
                       // FLAG information - store and evaluate
                       //------------------------------------------------------------------------------------------
                       // copy command setFlags for storing and usage in flag handling
                       // // setFlagsBuffer has twice the number of slots of PathDataPreBuffered to store flag information of past executed (already in MotionQueue) commands
                       #statFlagsBuffer.bufferElement[#statFlagsBuffer.writeBufferElement].pathDataName := #statPathDataPreBuffered.commands[#statPathDataPreBuffered.retrievePointer].pathDataName;
                       #statFlagsBuffer.bufferElement[#statFlagsBuffer.writeBufferElement].pathDataIdentifier := #statPathDataIdentifier;
                       #statFlagsBuffer.bufferElement[#statFlagsBuffer.writeBufferElement].cmdId := #statPathDataPreBuffered.commands[#statPathDataPreBuffered.retrievePointer].cmdID;
                       #statFlagsBuffer.bufferElement[#statFlagsBuffer.writeBufferElement].setFlags := #statPathDataPreBuffered.commands[#statPathDataPreBuffered.retrievePointer].setFlags;
                       #statFlagsBuffer.bufferElement[#statFlagsBuffer.writeBufferElement].valueFlags := #statPathDataPreBuffered.commands[#statPathDataPreBuffered.retrievePointer].valueFlags;
                       #statFlagsBuffer.bufferElement[#statFlagsBuffer.writeBufferElement].isIntermediateCmd := #statPathDataPreBuffered.commands[#statPathDataPreBuffered.retrievePointer].isIntermediateCmd;

                       // go to execution if cmd was copied
                       #statStateExecution := #EX_TRIGGERING_CMD;


                       IF #statPathDataPreBuffered.retrievePointer < "LKINCTRL_NO_OF_PATHDATA_PREBUFFER_ELEMENTS" THEN
                           #statPathDataPreBuffered.retrievePointer += 1;
                       ELSE
                           // restart PathDataPreBuf retrievePointer
                           #statPathDataPreBuffered.retrievePointer := 1;
                           // reset restart bit of pointer
                           #statPathDataPreBuffered.addPointerRestarted := FALSE;
                       END_IF;

                       #statSetFlagsBufferWriteBufferElement_old := #statFlagsBuffer.writeBufferElement;
                       // increase statSetFlagsBuffer write pointer and restart at overflow
                       IF #statFlagsBuffer.writeBufferElement < "LKINCTRL_NO_OF_SETFLAGS_BUFFER_ELEMENTS" THEN
                           #statFlagsBuffer.writeBufferElement := #statFlagsBuffer.writeBufferElement + 1;
                       ELSE
                           #statFlagsBuffer.writeBufferElement := 1;
                       END_IF;

                   ELSE
                       // set subfunction status according to PreBuffer status
                       IF (#statPathDataPreBuffered.retrievePointer = #statPathDataPreBuffered.addPointer
                           AND #statPathDataPreBuffered.addPointerRestarted = FALSE)
                       THEN
                           #statSubfunctionStatus := #STATUS_WAITING_FOR_PREBUFFERED_CMD;

                           // Check STOPRE signal from Parser/PreBuffer --> If true and executer is done then reset stopre to continue parsing
                           // PreBuffered commands are then executed and Parser and MovePath are in sync
                           IF #instLKinCtrl_MC_ExecuteKinMotionCmd.done AND #instLKinCtrl_PreBuffer.preprocessingStop THEN
                               #instLKinCtrl_PreBuffer.preprocessingStop := FALSE;
                           END_IF;


                       ELSIF (#statPathDataPreBuffered.addPointerRestarted = TRUE
                           AND (#statPathDataPreBuffered.retrievePointer - 1 = #statPathDataPreBuffered.addPointer))
                       THEN
                           #statSubfunctionStatus := #STATUS_PREBUFFERED_FULL;
                       END_IF;
                   END_IF;
                   // store old cmdID and PathDataName
                   #statPreBufferedCmdIdOld := #statPathDataElementPreBuffered.cmdID;
                   #statPreBufferedPathDataNameOld := #statPathDataElementPreBuffered.pathDataName;

                   // Check if interrupt was executed at start and if continue is needed
                   IF #statInterruptedAtStart THEN
                       IF #axesGroup.StatusMotionQueue.NumberOfCommands >= MIN(IN1:=#NO_OF_COMMANDS_PRELOADING, IN2:=#axesGroup.MotionQueue.MaxNumberOfCommands)
                           OR #statPathDataElementPreBuffered.cmdType = "LKINCTRL_CMD_WAIT_TIME" // Continue if waitTime shall be executed else we have deadlock
                           OR #statPathDataElementPreBuffered.cmdID = #statLastCmdIdPathdata // Continue if end of path was reached
                       THEN
                           #statStoreInterruptStateExecution := #statStateExecution;
                           #statStateExecution := #EX_CONTINUEING;
                           #statInterruptedAtStart := FALSE;
                       END_IF;
                   END_IF;

               END_IF;

           END_IF;
       END_REGION EX_GET_CMD


       // state reached when cmd should be triggered
       REGION EX_TRIGGERING_CMD
           IF #statStateExecution = #EX_TRIGGERING_CMD
               // AND #statDebugState = TRUE
               // wait condition bit (used for singleStep)
               AND #statExecutionWaitSingleStep = FALSE
               // wait condition bit (used for WAIT_TIME running)
               AND #statExecutionWaitTimerRunning = FALSE
               // wait condition bit (used for wait flags (acknowledge needed))
               AND #statWaitMain = FALSE
               // wait condition bit (used for wait value flags (acknowledge needed))
               AND #statWaitValueMain = FALSE
           THEN
               // reset  variable for single step debugging of states
               #statDebugState := FALSE;

               // call FB_ExecutePathMotion to execute cmd in same cycle
               #instLKinCtrl_MC_ExecuteKinMotionCmd(execute := TRUE,
                                                    interrupt := #interrupt,
                                                    stop := #stop,
                                                    pathDataElementPreBuf := #statPathDataElementPreBuffered,
                                                    conveyorConfiguration := #configuration.conveyorParameter,
                                                    to_Kinematics := #axesGroup);


               // check for cmd to be executed 
               IF #instLKinCtrl_MC_ExecuteKinMotionCmd.cmdExecuted THEN
                   // evaluate flag information for wait flags
                   // check for cmdId not to exceed array limits
                   IF #statFlagsBuffer.bufferElement[#statSetFlagsBufferWriteBufferElement_old].cmdId <> 0 THEN
                       // run through all setFlags in command
                       FOR #tempFlagCmdCounter := 1 TO "LKINCTRL_NO_OF_CMD_SETFLAGS" DO
                           // check preBuffered command for wait flag
                           IF #statFlagsBuffer.bufferElement[#statSetFlagsBufferWriteBufferElement_old].setFlags[#tempFlagCmdCounter].flag > -1
                               AND (#statFlagsBuffer.bufferElement[#statSetFlagsBufferWriteBufferElement_old].setFlags[#tempFlagCmdCounter].flagMode = 5
                               OR #statFlagsBuffer.bufferElement[#statSetFlagsBufferWriteBufferElement_old].setFlags[#tempFlagCmdCounter].flagMode = 15)
                           THEN
                               // increase counter to count activated wait flags in command
                               #statWaitFlags.waitCtr += 1;
                               // store information on which flags are wait flags
                               #statWaitFlags.waitFlag[#tempFlagCmdCounter] := #statFlagsBuffer.bufferElement[#statSetFlagsBufferWriteBufferElement_old].setFlags[#tempFlagCmdCounter].flag;
                           END_IF;
                       END_FOR;

                       // run through all valueFlags in command
                       FOR #tempFlagCmdCounter := 1 TO "LKINCTRL_NO_OF_CMD_VALUEFLAGS" DO
                           // check preBuffered command for wait flag
                           IF #statFlagsBuffer.bufferElement[#statSetFlagsBufferWriteBufferElement_old].valueFlags[#tempFlagCmdCounter].flag > -1
                               AND (#statFlagsBuffer.bufferElement[#statSetFlagsBufferWriteBufferElement_old].valueFlags[#tempFlagCmdCounter].flagMode = 5
                               OR #statFlagsBuffer.bufferElement[#statSetFlagsBufferWriteBufferElement_old].valueFlags[#tempFlagCmdCounter].flagMode = 15)
                           THEN
                               // increase counter to count activated wait value flags in command
                               #statWaitValueFlags.waitCtr += 1;
                               // store information on which flags are wait value flags
                               #statWaitValueFlags.waitFlag[#tempFlagCmdCounter] := #statFlagsBuffer.bufferElement[#statSetFlagsBufferWriteBufferElement_old].valueFlags[#tempFlagCmdCounter].flag;
                           END_IF;
                       END_FOR;
                   ELSE
                       // Do nothing, e.g. empty PathData element
                       ;
                   END_IF;

                   // go to state triggered when command has been successfully executed to MotionQueue
                   #statStateExecution := #EX_TRIGGERED_CMD;
               END_IF;

               // check for execution to be waiting for rising edge of execute to continue
           ELSIF (#statExecutionWaitSingleStep = TRUE
               OR #statWaitMain = TRUE
               OR #statWaitValueMain = TRUE
               OR #statExecutionWaitTimerRunning = TRUE)
               // check for no motion cmd to be active at TO_Kinematics
               AND #instLKinCtrl_MC_ExecuteKinMotionCmd.active = FALSE
               AND #statStateExecution = #EX_TRIGGERING_CMD // Added FR 2019/04/11
           THEN
               // set status accordingly
               #statStatus := #STATUS_EXECUTION_WAITING;
           END_IF;
       END_REGION EX_TRIGGERING_CMD


       // state reached when cmd has been triggered and is executed to the MotionQueue
       REGION EX_TRIGGERED_CMD
           IF #statStateExecution = #EX_TRIGGERED_CMD
               // AND #statDebugState = TRUE
           THEN
               // reset  variable for single step debugging of states
               #statDebugState := FALSE;

               // Overwrite status after ExecutionWaiting for correct flag behavior
               #statStatus := #STATUS_PATHMOTION_RUNNING; // Status is only active until StatusWord of kinematics overwrites it again

               // call FB_ExecutePathMotion to reset execute in same cycle after execution (for rising edge in next cycle)
               #instLKinCtrl_MC_ExecuteKinMotionCmd(execute := FALSE,
                                                    interrupt := #interrupt,
                                                    stop := #stop,
                                                    pathDataElementPreBuf := #statPathDataElementPreBuffered,
                                                    to_Kinematics := #axesGroup);

               // check for executed cmd to be last cmd in PathData
               IF #statPathDataElementPreBuffered.cmdID = #statLastCmdIdPathdata
                   AND #statPathDataElementPreBuffered.isIntermediateCmd = FALSE
               THEN
                   // go to state to wait for done / retriggering (no further cmds to be triggered)
                   #statStateExecution := #EX_ALL_TRIGGERED;
               ELSE
                   // go to EX_GET_CMD to get next command
                   #statStateExecution := #EX_GET_CMD;
               END_IF;


           END_IF;
       END_REGION EX_TRIGGERED_CMD


       // state reached when all cmds have been executed to the MotionQueue (wait for done or reTriggering)
       REGION EX_ALL_TRIGGERED
           IF #statStateExecution = #EX_ALL_TRIGGERED
               // AND #statDebugState = TRUE
           THEN
               // reset  variable for single step debugging of states
               #statDebugState := FALSE;

               // set status and status bit to set readyForNextPath output
               #statReadyForNextPath := TRUE;
               #statStatus := #STATUS_READYFORNEXTPATH;

               // Added remDistance check if no Motion Command follows after STOPRE --> Done signal is already false because it was checked in "GET_CMD"
               // wait for done signal of ExecuteKinMotionCmd (end of PathData reached)
               IF (#instLKinCtrl_MC_ExecuteKinMotionCmd.done
                   OR (#instLKinCtrl_MC_ExecuteKinMotionCmd.remainingDistanceActCmd = 0.0
                   AND #instLKinCtrl_MC_ExecuteKinMotionCmd.activeCmdNo = #statLastCmdIdPathdata
                   AND #instLKinCtrl_MC_ExecuteKinMotionCmd.active = FALSE
                   AND #instLKinCtrl_MC_ExecuteKinMotionCmd.busy = FALSE))
                   // no commmands in PathData ==> empty PathData
                   OR #statLastCmdIdPathdata = 0
                   // Executer was done but waitFlag was still active
                   OR #statExecuterWasDone
               THEN
                   // Wait until all setFlags and all valueFlags are acknowledged
                   IF NOT #statWaitMain AND NOT #statWaitValueMain THEN
                       // set status to set done output according to FB template
                       #statStatus := #STATUS_EXECUTION_FINISHED;
                       // Reset bit to memorize done output of MC_ExecuteKinMotionCmd
                       #statExecuterWasDone := FALSE;
                   ELSE
                       // Set status to waiting until all wait flags are acknowledged
                       #statStatus := #STATUS_EXECUTION_WAITING;
                       // Set bit to memorize done output of MC_ExecuteKinMotionCmd
                       #statExecuterWasDone := TRUE;
                   END_IF;
               END_IF;
           END_IF;
       END_REGION EX_TRIGGERED_CMD


       // state reached when GroupInterrupt is interrupted ==> do nothing when interrupted
       REGION EX_CONTINUEING
           IF #statStateExecution = #EX_CONTINUEING
               // AND #statDebugState = TRUE
           THEN
               // reset  variable for single step debugging of states
               #statDebugState := FALSE;

               // set continueMotion input on LKinCtrl_ExecuteKinMotionCmd
               #instLKinCtrl_MC_ExecuteKinMotionCmd.continueMotion := TRUE;

               // set state machine to CONTINUED after successfull continue of path motion
               IF #instLKinCtrl_MC_ExecuteKinMotionCmd.diagnostics.status = 16#7100 THEN
                   #statStateExecution := #EX_CONTINUED;
               END_IF;

           END_IF;
       END_REGION EX_CONTINUEING


       // state reached when GroupContinue is done ==> do nothing when path motion continues
       REGION EX_CONTINUED
           IF #statStateExecution = #EX_CONTINUED
               // AND #statDebugState = TRUE
           THEN
               // reset  variable for single step debugging of states
               #statDebugState := FALSE;

               // set status accordingly
               #statStatus := #STATUS_PATHMOTION_RUNNING;

               // reset continueMotion input on LKinCtrl_ExecuteKinMotionCmd
               #instLKinCtrl_MC_ExecuteKinMotionCmd.continueMotion := FALSE;

               // reset state machine to state before interrupt
               #statStateExecution := #statStoreInterruptStateExecution;

           END_IF;
       END_REGION EX_CONTINUED

       // state reached to execute MC_GroupInterrupt ==> wait for interrupt to be done
       REGION EX_INTERRUPTING
           IF #statStateExecution = #EX_INTERRUPTING
               // AND #statDebugState = TRUE
           THEN
               // reset  variable for single step debugging of states
               #statDebugState := FALSE;

               // reset trigger for cmd execution at LKinCtrl_ExecuteKinMotionCmd to enable new rising edge after continue
               // FR 11.03.2020: do not reset execute when wait time is running to avoid triggering the same time twice
               IF NOT #statExecutionWaitTimerRunning THEN
                   #instLKinCtrl_MC_ExecuteKinMotionCmd.execute := FALSE;
               END_IF;
               #instLKinCtrl_MC_ExecuteKinMotionCmd.continueMotion := FALSE; // FR 11.03.2020: Also reset continue input

               // check for path motion to have been interrupted (by LKinCtrlExecuteKinMotionCmd)
               IF #instLKinCtrl_MC_ExecuteKinMotionCmd.diagnostics.status = 16#7102 THEN
                   #statStateExecution := #EX_INTERRUPTED;
               END_IF;

           END_IF;
       END_REGION EX_INTERRUPTING


       // state reached when path motion has been interrupted in LKinExectuteKinMotionCmd
       REGION EX_INTERRUPTED
           IF #statStateExecution = #EX_INTERRUPTED
               // AND #statDebugState = TRUE
           THEN
               // reset  variable for single step debugging of states
               #statDebugState := FALSE;

               // set status accordingly
               #statStatus := #STATUS_PATHMOTION_INTERRUPTED;

               // do nothing, wait in this state

           END_IF;
       END_REGION EX_INTERRUPTED

       // state reached when stop input is triggered (path motion stop is executed in LKinExectuteKinMotionCmd)
       REGION EX_STOPPING
           IF #statStateExecution = #EX_STOPPING
               // AND #statDebugState = TRUE
           THEN
               // reset variable for single step debugging of states
               #statDebugState := FALSE;

               // set status accordingly
               #statStatus := #STATUS_PATHMOTION_STOPPING;

               // check for path motion to be aborted in LKinExectuteKinMotionCmd
               IF #instLKinCtrl_MC_ExecuteKinMotionCmd.commandAborted THEN
                   #statStateExecution := #EX_STOPPED_STATE;

               ELSIF #instLKinCtrl_MC_ExecuteKinMotionCmd.diagnostics.status.%X15 THEN // check for executer status >= 16#8000
                   #statStateExecution := #EX_ERROR_STATE;
                   #statStatus := #ERR_EXECUTE_KINMOTIONCMD;
                   #statSubfunctionStatus := #instLKinCtrl_MC_ExecuteKinMotionCmd.diagnostics.status;
               END_IF;

           END_IF;
       END_REGION EX_STOPPING


       // state reached when path motion has been stopped in LKinExectuteKinMotionCmd
       REGION EX_STOPPED_STATE
           IF #statStateExecution = #EX_STOPPED_STATE
               // AND #statDebugState = TRUE
           THEN
               // reset  variable for single step debugging of states
               #statDebugState := FALSE;

               // set status accordingly
               #statStatus := #STATUS_COMMAND_ABORTED;
               #statSubfunctionStatus := #instLKinCtrl_MC_ExecuteKinMotionCmd.diagnostics.status;

               //------------------------------------------------------------------------------------------
               // added 2020.02.07 DF: call Prebuffer with false (reset retrievePointer)
               #instLKinCtrl_PreBuffer(enable := FALSE,
                                       to_Kinematics := #axesGroup,
                                       pathData := #pathData,
                                       pathDataPreBuf := #statPathDataPreBuffered);
               //------------------------------------------------------------------------------------------
               // do nothing, wait in this state

           END_IF;
       END_REGION EX_STOPPED_STATE


       // state reached when error occured ==> do nothing when error occured
       REGION EX_ERROR_STATE
           IF #statStateExecution = #EX_ERROR_STATE
               // AND #statDebugState = TRUE
           THEN
               // reset  variable for single step debugging of states
               #statDebugState := FALSE;

               IF #instLKinCtrl_PreBuffer.error THEN
                   IF #axesGroup.StatusPath.Velocity = 0.0                     // TO Kinematics velocity 0.0
                       AND #axesGroup.StatusWord.%X12                            // TO Kinematics in constant velocity
                       AND #axesGroup.StatusMotionQueue.NumberOfCommands = 0     // all commands deleted from MotionQueue
                   THEN
                       // do nothing if path motion has already been stopped, no stop execution necessary
                       ;
                   ELSE
                       // trigger #stop at LKinCtrl_ExecuteKinMotionCmd in case of #error in #pathData and path already running
                       #tempStop := TRUE;
                   END_IF;
               END_IF;

               // store LKinCtrl_ExecuteKinMotionCmd error before resetting trigger
               IF #instLKinCtrl_MC_ExecuteKinMotionCmd.error THEN
                   #statSubfunctionStatus := #instLKinCtrl_MC_ExecuteKinMotionCmd.diagnostics.status;
               END_IF;

               IF (#statStatus = #STATUS_STOP_DUE_TO_ERROR AND #instLKinCtrl_MC_ExecuteKinMotionCmd.commandAborted)
                   OR (#tempStop AND #instLKinCtrl_MC_ExecuteKinMotionCmd.error) // Check if stop also failed with error
               THEN
                   #statStatus := #ERR_EXECUTE_KINMOTIONCMD;
               END_IF;

               // Set stop to true
               IF #statStatus = #STATUS_STOP_DUE_TO_ERROR THEN
                   #tempStop := TRUE;
               END_IF;

               // reset trigger for FB LKinExecuteKinMotionCmd
               #instLKinCtrl_MC_ExecuteKinMotionCmd.execute := FALSE;
           END_IF;

       END_REGION EX_ERROR_STATE

   END_REGION EXECUTION


   REGION CALL_FB_EXECUTE
       // call FB LKinCtrl_ExecuteKinMotionCmd in every cycle to keep FB outputs updated
       #instLKinCtrl_MC_ExecuteKinMotionCmd(interrupt := #tempInterrupt AND #statDone = FALSE, // If done then interrupting leads to trouble
                                            stop := #tempStop,
                                            stopMode := #configuration.stopMode,
                                            writtenActiveCmdNo := #statWrittenActiveCmdNo,
                                            waitTimeActive => #statExecutionWaitTimerRunning,
                                            pathDataElementPreBuf := #statPathDataElementPreBuffered,
                                            to_Kinematics := #axesGroup);

       // FR 18.03.2020: Check done bit here for correct timing of active, busy & done
       // wait for done signal of ExecuteKinMotionCmd (end of PathData reached)
       IF #statStateExecution = #EX_ALL_TRIGGERED
           AND (#instLKinCtrl_MC_ExecuteKinMotionCmd.done
           // no commmands in PathData ==> empty PathData
           OR #statLastCmdIdPathdata = 0
           // Executer was done but waitFlag was still active
           OR #statExecuterWasDone)
       THEN
           // Wait until all setFlags are acknowledged
           IF NOT #statWaitMain
               // also wait until all valueFlags
               AND NOT #statWaitValueMain
           THEN
               // set status to set done output according to FB template
               #statStatus := #STATUS_EXECUTION_FINISHED;

               // Reset bit to memorize done output of MC_ExecuteKinMotionCmd
               #statExecuterWasDone := FALSE;
           ELSE
               // Set status to waiting until all wait flags are acknowledged
               #statStatus := #STATUS_EXECUTION_WAITING;

               // Set bit to memorize done output of MC_ExecuteKinMotionCmd
               #statExecuterWasDone := TRUE;
           END_IF;
       END_IF;

       // detect error in path execution in FB LKinCtrl_ExecuteKinMotionCmd
       IF #instLKinCtrl_MC_ExecuteKinMotionCmd.error THEN
           // set status accordingly
           IF #instLKinCtrl_MC_ExecuteKinMotionCmd.diagnostics.status = 16#8245 // Error at Kinematics --> Nothing more to do
               OR #instLKinCtrl_MC_ExecuteKinMotionCmd.diagnostics.status = 16#8244 THEN // Error GroupStop failed --> Nothing more to do
               #statStatus := #ERR_EXECUTE_KINMOTIONCMD;
           ELSE
               #statStatus := #STATUS_STOP_DUE_TO_ERROR; // Error at command --> Stop Kinematics
           END_IF;

           #statSubfunctionStatus := #instLKinCtrl_MC_ExecuteKinMotionCmd.diagnostics.status;

           // set state machine to error state
           #statStateExecution := #EX_ERROR_STATE;

       END_IF;

       // detect stopping to be in progress (here external stop, internal handled immediately)
       IF #instLKinCtrl_MC_ExecuteKinMotionCmd.diagnostics.status = 16#7103 // Executer is stopping
           // do not go to stopping state and overwrite status when PreBuffer detected error first
           AND #instLKinCtrl_PreBuffer.error = FALSE
           AND #statStatus <> #STATUS_STOP_DUE_TO_ERROR
       THEN
           // set status accordingly
           #statStateExecution := #EX_STOPPING;
           #statSubfunctionStatus := #instLKinCtrl_MC_ExecuteKinMotionCmd.diagnostics.status;
       END_IF;

   END_REGION CALL_FB_EXECUTE


   REGION STATIC_VARIABLE_HANDLING


       // set status in case no specific status has been set before
       IF #statStatus.%X15 = FALSE                                                 // no error deteceted
           AND #statStatus <> #STATUS_COMMAND_ABORTED                                  // no abort/stop detected
           AND #statStatus <> #STATUS_PATHMOTION_INTERRUPTED                           // no interrupt deteceted
           AND #statStatus <> #STATUS_EXECUTION_FINISHED                               // no completion of path motion detected
           AND #statStatus <> #STATUS_READYFORNEXTPATH                                 // no readyForNextPath signalized
           AND #statStatus <> #STATUS_NO_CALL                                          // fb not about to be deactivated in next cycle
           AND #statStatus <> #STATUS_PATHMOTION_STOPPING                              // no stopping in progress detected
           AND #statStatus <> #STATUS_STOP_DUE_TO_ERROR
       THEN
           // check for linear command to be active 
           IF #axesGroup.StatusWord.%X8 THEN
               #statStatus := #STATUS_CMD_LIN_ACTIVE;

               // check for circulat command to be active
           ELSIF #axesGroup.StatusWord.%X9 THEN
               #statStatus := #STATUS_CMD_CIRC_ACTIVE;

               // check for move direct command to be active
           ELSIF #axesGroup.StatusWord.%X11 THEN
               #statStatus := #STATUS_CMD_MOVE_DIRECT_ACTIVE;

               // Check for waitTimerRunning
           ELSIF #statExecutionWaitTimerRunning THEN
               #statStatus := #STATUS_EXECUTION_WAITING;
           END_IF;
       END_IF;


   END_REGION


   REGION OUTPUTS

       REGION FLAG_HANDLING
           // Call FlagHandling FBs
           //------------------------------------------------------------------------------------------
           // FR 16.03.2020: Reworked Flag FBs
           // Enable flag FBs when not finished and not no call (resetting)
           IF #statStatus <> #STATUS_EXECUTION_FINISHED AND #statStatus <> #STATUS_NO_CALL THEN
               #instLKinCtrl_SetFlagCtrl.enable := TRUE;
               #instLKinCtrl_ValueFlagCtrl.enable := TRUE;
           ELSE
               #instLKinCtrl_SetFlagCtrl.enable := FALSE;
               #instLKinCtrl_ValueFlagCtrl.enable := FALSE;
           END_IF;

           // Boolean Flags
           #instLKinCtrl_SetFlagCtrl(activeCmdNo := #instLKinCtrl_MC_ExecuteKinMotionCmd.activeCmdNo,
                                     activePathDataIdentifier := #instLKinCtrl_MC_ExecuteKinMotionCmd.activePathDataIdentifier,
                                     activePathDataName := #instLKinCtrl_MC_ExecuteKinMotionCmd.activePathDataName,
                                     remainingDistanceActCmd := #instLKinCtrl_MC_ExecuteKinMotionCmd.remainingDistanceActCmd,
                                     kinematicsStatusWord := #axesGroup.StatusWord,
                                     movePathStatus := #statStatus,
                                     flagsBuffer := #statFlagsBuffer,
                                     waitMain => #statWaitMain,
                                     flags := #flags,
                                     waitFlags := #statWaitFlags);

           // Check if flag control FB has thrown an error
           IF #instLKinCtrl_SetFlagCtrl.error THEN
               #statStatus := #ERR_SET_FLAG_CONTROL;
               #statSubfunctionStatus := #instLKinCtrl_SetFlagCtrl.status;
           END_IF;


           // LReal Flags
           #instLKinCtrl_ValueFlagCtrl(activeCmdNo := #instLKinCtrl_MC_ExecuteKinMotionCmd.activeCmdNo,
                                       activePathDataIdentifier := #instLKinCtrl_MC_ExecuteKinMotionCmd.activePathDataIdentifier,
                                       activePathDataName := #instLKinCtrl_MC_ExecuteKinMotionCmd.activePathDataName,
                                       remainingDistanceActCmd := #instLKinCtrl_MC_ExecuteKinMotionCmd.remainingDistanceActCmd,
                                       kinematicsStatusWord := #axesGroup.StatusWord,
                                       movePathStatus := #statStatus,
                                       flagsBuffer := #statFlagsBuffer,
                                       waitMain => #statWaitValueMain,
                                       valueFlags := #valueFlags,
                                       waitFlags := #statWaitValueFlags);

           // Check if flag control FB has thrown an error
           IF #instLKinCtrl_ValueFlagCtrl.error THEN
               #statStatus := #ERR_VALUE_FLAG_CONTROL;
               #statSubfunctionStatus := #instLKinCtrl_ValueFlagCtrl.status;
           END_IF;

           // Save written active cmd number for "ExecuteKinMotionCmd" input
           #statWrittenActiveCmdNo := #instLKinCtrl_MC_ExecuteKinMotionCmd.activeCmdNo;
       END_REGION FLAG_HANDLING


       REGION STATUS_EVALUATION
           // Write outputs
           IF (#statStatus = #STATUS_EXECUTION_FINISHED) AND (#statDone = FALSE) THEN // Execution finished without errors
               #statDone := TRUE;
               #statBusy := FALSE;
               #statCommandAborted := FALSE;
               #statError := FALSE;
               #statStateExecution := #EX_NO_PROCESSING; // Switch state machine to "no processing"

           ELSIF (#statStatus.%X15 = TRUE) AND (#statError = FALSE) THEN // Error occurred (#statStatus is 16#8000 to 16#FFFF)
               #statDone := FALSE;
               #statBusy := FALSE;
               #statCommandAborted := FALSE;
               #statError := TRUE;
               // Write diagnostics
               #diagnostics.stateMovePath := #statStateExecution;
               #status := #statStatus;
               #diagnostics.statusSubFunction := #statSubfunctionStatus;
               #statStateExecution := #EX_ERROR_STATE; // Switch state machine to "no processing"

           ELSIF (#statStatus = #STATUS_COMMAND_ABORTED) AND (#statCommandAborted = FALSE) THEN // Commanded functionality has been aborted by another command
               #statDone := FALSE;
               #statBusy := FALSE;
               #statCommandAborted := TRUE;
               #statError := FALSE;
               // Write diagnostics
               #diagnostics.stateMovePath := #statStateExecution;
               #status := #statStatus;
               #diagnostics.statusSubFunction := #statSubfunctionStatus;
               #statStateExecution := #EX_NO_PROCESSING; // Switch state machine to "no processing"

           ELSIF (#tempExecute = FALSE) AND (#tempStop = FALSE) AND ((#statDone = TRUE) OR (#statError = TRUE) OR (#statCommandAborted = TRUE)) THEN // Reset outputs
               #statDone := FALSE;
               #statBusy := FALSE;
               #statCommandAborted := FALSE;
               #statError := FALSE;
               #statReadyForNextPath := TRUE; // Added FR 2019/04/11
               #statStatus := #STATUS_NO_CALL;
           END_IF;

           // Write static values to outputs
           #done := #statDone;
           #busy := #statBusy;
           #active := #instLKinCtrl_MC_ExecuteKinMotionCmd.active;
           #commandAborted := #statCommandAborted;
           #error := #statError;
           // check for error to be pending
           IF #statError THEN
               // write status to errorID in case of error pending
               #statErrorID := #statStatus;
           ELSE
               // do nothing
               ;
           END_IF;
           #diagnostics.errorID := #statErrorID;
           #status := #statStatus;
           #diagnostics.stateMovePath := #statStateExecution;
           // write diagnostics information according to pending error type
           IF #instLKinCtrl_PreBuffer.error = FALSE THEN
               // write usual data to outputs
               #diagnostics.motionFBStatus := #instLKinCtrl_MC_ExecuteKinMotionCmd.diagnostics.motionFBstatus;
               #diagnostics.motionFBNumber := #instLKinCtrl_MC_ExecuteKinMotionCmd.diagnostics.faultFBNumber;
               #diagnostics.pathDataName := #instLKinCtrl_MC_ExecuteKinMotionCmd.diagnostics.faultPathDataName;
               #diagnostics.cmdNumber := #instLKinCtrl_MC_ExecuteKinMotionCmd.diagnostics.faultSetNumber;
               #diagnostics.kinematicsErrorWord := #instLKinCtrl_MC_ExecuteKinMotionCmd.diagnostics.kinematicsErrorWord;
           ELSE
               // write error specific data to outputs in case of wrong PathData parametrization
               #diagnostics.motionFBStatus := #instLKinCtrl_PreBuffer.status;
               #diagnostics.pathDataName := #statPathDataPreBuffered.pathDataName;
               #diagnostics.cmdNumber := #instLKinCtrl_PreBuffer.pathDataRetrievePointer;
           END_IF;

           #diagnostics.kinematicsStatusWord := #instLKinCtrl_MC_ExecuteKinMotionCmd.diagnostics.kinematicsStatusWord;
           #activePathData := #instLKinCtrl_MC_ExecuteKinMotionCmd.activePathDataName;
           #activeCmdNo := #instLKinCtrl_MC_ExecuteKinMotionCmd.activeCmdNo;
           #remainingDistanceActCmd := #instLKinCtrl_MC_ExecuteKinMotionCmd.remainingDistanceActCmd;
           #readyForNextPath := #statReadyForNextPath;

       END_REGION STATUS_EVALUATION

   END_REGION OUTPUTS

   // =================================================================================================================
   // End of Function Block: LKinCtrl_MC_MovePath
   // =================================================================================================================
END_FUNCTION_BLOCK

FUNCTION_BLOCK "LKinCtrl_MC_JogFrame"   // FB35010, SCL
TITLE = LKinCtrl_MC_JogFrame
{ S7_Optimized_Access := 'TRUE' }
AUTHOR : tech.team.motioncontrol@siemens.com
FAMILY : LKinCtrl
VERSION : 1.1
// Functionality: This function block provides various jog functionality for kinematics technology object.
   VAR_INPUT
      jogForward : Bool := FALSE;   // Jog the kinematics forward in the selected jog direction
      jogBackward : Bool := FALSE;   // Jog the kinematics backward in the selected jog direction
      jogToPosition : Bool := FALSE;   // Jog the kinematics to the specified target position
      jogDirection : USInt := 1;   // 1=x-direction, 2=y-direction, 3=z-direction, 4=a-direction
      jogModeInc : Bool := FALSE;   // 1=incremental jog mode, 0=continuous jog mode
      jogIncrement : LReal := 1.0;   // Specification of the jog increment
      targetPosition : "LKinCtrl_typeCartesianPosition";   // Specification of the target position
      coordSystem : DInt := 0;   // 0=WCS, 1= OCS1, 2=OCS2, 3=OCS3
      tool : DInt := 1;   // 1= tool1, 2=tool2, 3=tool3
      dynamics : "LKinCtrl_typeDynamics";   // Specification of the jog dynamics
   END_VAR
   VAR_OUTPUT
      done : Bool := FALSE;   // TRUE: Commanded functionality has been completed successfully
      busy : Bool := FALSE;   // TRUE: FB is not finished and new output values can be expected
      active : Bool := FALSE;   // TRUE: The setpoints are calculated
      error : Bool := FALSE;   // TRUE: An error occurred during the execution of the FB
      status : Word := 16#7000;   // 16#0000 - 16#7FFF: Status of the FB, 16#8000 - 16#FFFF: Error identification
      remainingDistance : LReal := 0.0;   // Distance-to-go of the current job
      diagnostics : "LKinCtrl_typeJogFrameDiagnostics";   // Diagnostics information
   END_VAR
   VAR_IN_OUT
      axesGroup : TO_Kinematics;   // Kinematics technology object
   END_VAR
   VAR
      instMC_SetTool : MC_SETTOOL;   // Instance MC_SetTool
      instMC_GroupStop : MC_GROUPSTOP;   // Instance MC_GroupStop
      instMC_MoveLinearAbsoute : MC_MOVELINEARABSOLUTE;   // Instance MC_MoveLinearAbsolute
      instMC_MoveLinearRelative : MC_MOVELINEARRELATIVE;   // Instance MC_MoveLinearRelative
      statDone : Bool := FALSE;   // Static value for output 'done'
      statBusy : Bool := FALSE;   // Static value for output 'busy'
      statActive : Bool := FALSE;   // Static value for output 'active'
      statError : Bool := FALSE;   // Static value for output 'error'
      statStatus : Word := 16#7000;   // 0000=STATUS_EXECUTION_FINISHED; 7000=STATUS_NO_CALL; 7001=STATUS_FIRST_CALL; 7002=STATUS_SUBSEQUENT_CALL; 8600=ERR_UNDEFINED_STATE
      statRemainingDistance : LReal := 0.0;   // Static value for remaining distance
      statFBState : DInt := 0;   // 0= NO PROCESSING; 10=IDLE; 20=SET_TOOL; 30=SET_DYNAMICS, 50=EXECUTE_MOVEMENT; 100=STOP
      statToolOld : DInt := 1;   // Static value for tool
      statJogForwardOld : Bool := FALSE;   // Static value for jog forward command
      statJogBackwardOld : Bool := FALSE;   // Static value for jog backward command
      statJogToPositionOld : Bool := FALSE;   // Static value for jog to position command
      statOrientationDynamicsChanged : Bool := FALSE;   // Static value indicates that default orientation dynamics have been changed
      statOrientationDynamicsOld : "LKinCtrl_typePathDynamics";   // Static value for orientation dynamics
   END_VAR
   VAR_TEMP
      tempJogForward : Bool;   // Temporary variable for jog forward input
      tempJogBackward : Bool;   // Temporary variable for jog backward input
      tempJogToPosition : Bool;   // Temporary variable for jog to position input
      tempCounter : DInt;   // Temporary variable for counter
      tempRet : Int;   // Temporary variable for time stamp if error occurred
   END_VAR
   VAR CONSTANT
      FB_STATE_NO_PROCESSING : DInt := 0;   // FB state: No processing
      FB_STATE_CMD_CONFIGURATION : DInt := 10;   // FB state: Basic command configuration are set depending on input parameter
      FB_STATE_SET_TOOL : DInt := 20;   // FB state: Tool change is performed if required
      FB_STATE_SET_DYNAMICS : DInt := 30;   // FB state: Dynamics configuration for jog command
      FB_STATE_EXECUTE_MOVEMENT : DInt := 50;   // FB state: Command is being executed
      FB_STATE_STOP : DInt := 100;   // FB state: Kinematics movement is stopped
      STATUS_EXECUTION_FINISHED : Word := 16#0000;   // The command execution is finished by reaching the target position or stopping the jog command
      STATUS_NO_CALL : Word := 16#7000;   // No call of FB
      STATUS_FIRST_CALL : Word := 16#7001;   // First cycle of FB after enabling
      STATUS_SUBSEQUENT_CALL : Word := 16#7002;   // FB enabled
      ERR_UNDEFINED_STATE : Word := 16#8600;   // Error due to an undefined FB state
      ERR_TO_KINEMATICS : Word := 16#8001;   // Error at technology object kinematics
      ERR_INVALID_JOG_DIRECTION : Word := 16#8007;   // The specified jog direction is invalid (valid values are 1=x-direction, 2=y-direction, 3=z-direction, 4=a-direction)
      ERR_MOTION_JOB_IN_PROGRESS : Word := 16#8090;   // A motion job is in progress or the kinematics control panel is activated
      ERR_TWO_JOG_COMMANDS_SIMULTANEOUSLY : Word := 16#8091;   // Two jog commands were triggered simultaneously
      ERR_INVALID_COORDINATE_SYSTEM : Word := 16#80B1;   // The specified coordinate system is invalid (valid values are 0=WCS, 1= OCS1, 2=OCS2, 3=OCS3)
      ERR_INVALID_TOOL : Word := 16#80CA;   // The specified tool is invalid (valid values are 1= tool1, 2=tool2, 3=tool3)
      MAX_DISTANCE : LReal := 700000000000.0;   // The value is set for relative linear movement as jog increment for icremental jog mode
      L_BOUND_TOOL : DInt := 1;   // Lower bound for tool selection
      U_BOUND_TOOL : DInt := 3;   // Upper bound for tool selection
      L_BOUND_JOG_DIRECTION : DInt := 1;   // Lower bound for jog direction selection
      U_BOUND_JOG_DIRECTION : DInt := 4;   // Upper bound for jog direction selection
      L_BOUND_COORDSYSTEM : DInt := 0;   // Lower bound for coordinate system selection
      U_BOUND_COORDSYSTEM : DInt := 3;   // Upper bound for coordinate system selection
   END_VAR
BEGIN
   //=============================================================================
   // SIEMENS AG
   // (c)Copyright 2018 All Rights Reserved
   //-----------------------------------------------------------------------------
   // Library:       LKinCtrl
   // Tested with:   S7-1516T
   // Engineering:   TIA Portal V15
   // Restrictions:  -
   // Requirements:  S7-1500T FW 2.5
   // Functionality: LKinCtrl_MC_JogFrame
   // This function block provides various jog functionality for kinematics technology object
   // 
   // Support: tech.team.motioncontrol@siemens.com
   // Note: Parameter comments are only available in language 'English (United States)'
   //-----------------------------------------------------------------------------
   // Change log table:
   // Version  Date        Expert in charge   Changes applied
   // 01.00.00 05.04.2018  IP                 First released version
   // 01.00.01 24.04.2018  IP                 Hotfix - initialization - no functional changes
   // 01.01.00 31.07.2018  IP                 Adjustment of input validation
   //                                         New wait condition for next movement until stopping is done
   //                                         Additional output parameter active and remaining distance
   // 01.01.01 07.08.2018  IP                 Hotfix - constant MAX_DISTANCE decreased
   // 01.01.02 09.01.2019  IP                 Hotfix - error indification adjusted
   // 01.01.03 14.01.2019  IP                 Hotfix - dynamics configuration adjusted
   //=============================================================================

   #tempJogForward := #jogForward; // Work with temporary value / create process image
   #tempJogBackward := #jogBackward;
   #tempJogToPosition := #jogToPosition;

   REGION TRIGGERING

     IF ((#tempJogForward AND NOT #statJogForwardOld) // Check if FB is triggered
       OR (#tempJogBackward AND NOT #statJogBackwardOld)
       OR (#tempJogToPosition AND NOT #statJogToPositionOld))
       AND (#statStatus = #STATUS_NO_CALL)
       AND (#statFBState = #FB_STATE_NO_PROCESSING)
     THEN

       // First call; set FB variables for outputs
       #statBusy := TRUE;
       #statDone := FALSE;
       #statActive := FALSE;
       #statError := FALSE;
       #statRemainingDistance := 0.0;
       #statStatus := #STATUS_FIRST_CALL;

       // check if input parameter are valid
       IF (#jogDirection < #L_BOUND_JOG_DIRECTION OR #jogDirection > #U_BOUND_JOG_DIRECTION) // check jog direction
         AND NOT #tempJogToPosition THEN
         #statStatus := #ERR_INVALID_JOG_DIRECTION;
       ELSIF #tool < #L_BOUND_TOOL OR #tool > #U_BOUND_TOOL THEN // check tool
         #statStatus := #ERR_INVALID_TOOL;
       ELSIF #coordSystem < #L_BOUND_COORDSYSTEM OR #coordSystem > #U_BOUND_COORDSYSTEM THEN // check coordinate system
         #statStatus := #ERR_INVALID_COORDINATE_SYSTEM;
       ELSIF NOT #axesGroup.StatusWord.%X6 THEN // check if a motion job is in progress or the kinematics control panel is activated
         #statStatus := #ERR_MOTION_JOB_IN_PROGRESS;
       ELSE // all input parameter are valid

         // reset execute inputs
         #instMC_GroupStop.Execute := FALSE;
         #instMC_MoveLinearAbsoute.Execute := FALSE;
         #instMC_MoveLinearRelative.Execute := FALSE;
         #instMC_SetTool.Execute := FALSE;

         // call FBs with execute = false
         #instMC_GroupStop(AxesGroup := #axesGroup);
         #instMC_MoveLinearAbsoute(AxesGroup := #axesGroup);
         #instMC_MoveLinearRelative(AxesGroup := #axesGroup);
         #instMC_SetTool(AxesGroup := #axesGroup);

         // get actual tool number
         #statToolOld := #axesGroup.StatusTool.ActiveTool;

         // safe default dynimcs for orientation axis
         #statOrientationDynamicsOld.velocity := #axesGroup.DynamicDefaults.Orientation.Velocity;
         #statOrientationDynamicsOld.acceleration := #axesGroup.DynamicDefaults.Orientation.Acceleration;
         #statOrientationDynamicsOld.deceleration := #axesGroup.DynamicDefaults.Orientation.Deceleration;
         #statOrientationDynamicsOld.jerk := #axesGroup.DynamicDefaults.Orientation.Jerk;
         #statOrientationDynamicsChanged := FALSE;

         // state machine - start functionality
         #statFBState := #FB_STATE_CMD_CONFIGURATION;
       END_IF;

     ELSIF (#statStatus = #STATUS_FIRST_CALL) THEN
       #statStatus := #STATUS_SUBSEQUENT_CALL;
     END_IF;

   END_REGION TRIGGERING

   IF (#statStatus = #STATUS_NO_CALL) THEN // Nothing to do -> End here to reduce "system load"
     RETURN;
   END_IF;

   REGION STOP_MOTION

     // detection of falling edge on jog command
     IF ((NOT #tempJogForward AND #statJogForwardOld)
       OR (NOT #tempJogBackward AND #statJogBackwardOld)
       OR (NOT #tempJogToPosition AND #statJogToPositionOld))
       AND NOT (#statFBState = #FB_STATE_NO_PROCESSING)
     THEN // stop jog command
       #statFBState := #FB_STATE_STOP;

       // two jog commands simultaneously    
     ELSIF ((#tempJogBackward AND #tempJogForward)
       OR (#tempJogBackward AND #tempJogToPosition)
       OR (#tempJogForward AND #tempJogToPosition))
       AND NOT (#statFBState = #FB_STATE_NO_PROCESSING)
     THEN // stop jog command
       #statFBState := #FB_STATE_STOP;
       #statStatus := #ERR_TWO_JOG_COMMANDS_SIMULTANEOUSLY;
     END_IF;

     IF #statStatus <> #STATUS_FIRST_CALL AND (#statStatus.%X15 = FALSE) THEN
       IF #axesGroup.StatusWord.%X1 // general TO error
         OR #instMC_MoveLinearRelative.Error
         OR #instMC_GroupStop.Error
         OR #instMC_MoveLinearAbsoute.Error
         OR #instMC_SetTool.Error
       THEN
         #statFBState := #FB_STATE_STOP;
       END_IF;
     END_IF;

   END_REGION

   // Edge detection 'execute' input
   #statJogForwardOld := #tempJogForward;
   #statJogBackwardOld := #tempJogBackward;
   #statJogToPositionOld := #tempJogToPosition;

   REGION RESET_DEFAULT_ORIENTATION_DYNAMICS

     IF (#instMC_MoveLinearRelative.Busy OR #instMC_MoveLinearAbsoute.Busy OR #statFBState = #FB_STATE_STOP)
       AND #statOrientationDynamicsChanged
     THEN // reset default orientation dynamics
       #axesGroup.DynamicDefaults.Orientation.Velocity := #statOrientationDynamicsOld.velocity;
       #axesGroup.DynamicDefaults.Orientation.Acceleration := #statOrientationDynamicsOld.acceleration;
       #axesGroup.DynamicDefaults.Orientation.Deceleration := #statOrientationDynamicsOld.deceleration;
       #axesGroup.DynamicDefaults.Orientation.Jerk := #statOrientationDynamicsOld.jerk;
       #statOrientationDynamicsChanged := FALSE;
     END_IF;

   END_REGION

   REGION ACTIVE_OUTPUT

     // set active output if any of motion commands is active
     IF #instMC_MoveLinearAbsoute.Active OR #instMC_MoveLinearRelative.Active OR #instMC_GroupStop.Active THEN
       #statActive := TRUE;
     ELSE
       #statActive := FALSE;
     END_IF;

   END_REGION

   REGION REMAINING_DISTANCE

     // set remaining distance at output if incremental mode active or while jogging to target position
     IF #instMC_MoveLinearAbsoute.Busy THEN
       #statRemainingDistance := #instMC_MoveLinearAbsoute.RemainingDistance;
     ELSIF #instMC_MoveLinearRelative.Busy AND #jogModeInc THEN
       #statRemainingDistance := #instMC_MoveLinearRelative.RemainingDistance;
     ELSE
       #statRemainingDistance := 0.0;
     END_IF;

   END_REGION

   REGION STATE_MACHINE

     CASE #statFBState OF // State machine of FB
       #FB_STATE_NO_PROCESSING: // No processing active (Note: this state must always be present and left empty)
         ;

       #FB_STATE_CMD_CONFIGURATION:

         REGION CONFIGURATION

           // jog forward or backward
           //*********************************************************************************************************
           IF #tempJogForward OR #tempJogBackward THEN
             // set MC_MoveLinearRelative parameter
             #instMC_MoveLinearRelative.CoordSystem := #coordSystem;
             #instMC_MoveLinearRelative.Velocity := #dynamics.path.velocity;
             #instMC_MoveLinearRelative.Acceleration := #dynamics.path.acceleration;
             #instMC_MoveLinearRelative.Deceleration := #dynamics.path.deceleration;
             #instMC_MoveLinearRelative.Jerk := #dynamics.path.jerk;

             // initialize jog distance - clear old values
             FOR #tempCounter := 1 TO 4 DO
               #instMC_MoveLinearRelative.Distance[#tempCounter] := 0.0;
             END_FOR;

             // set jog mode
             IF #jogModeInc THEN // incremental
               IF #tempJogForward THEN
                 #instMC_MoveLinearRelative.Distance[#jogDirection] := #jogIncrement;
               ELSIF #tempJogBackward THEN
                 #instMC_MoveLinearRelative.Distance[#jogDirection] := - #jogIncrement;
               END_IF;
               #instMC_MoveLinearRelative.DynamicAdaption := #dynamics.dynamicAdaption;

             ELSE // continouos
               IF #tempJogForward THEN
                 #instMC_MoveLinearRelative.Distance[#jogDirection] := #MAX_DISTANCE;
               ELSIF #tempJogBackward THEN
                 #instMC_MoveLinearRelative.Distance[#jogDirection] := - #MAX_DISTANCE;
               END_IF;

               // switch off dynamic adaption for continouos mode
               #instMC_MoveLinearRelative.DynamicAdaption := 0;
             END_IF;

